REGION Network 9: Mapare elemente safety
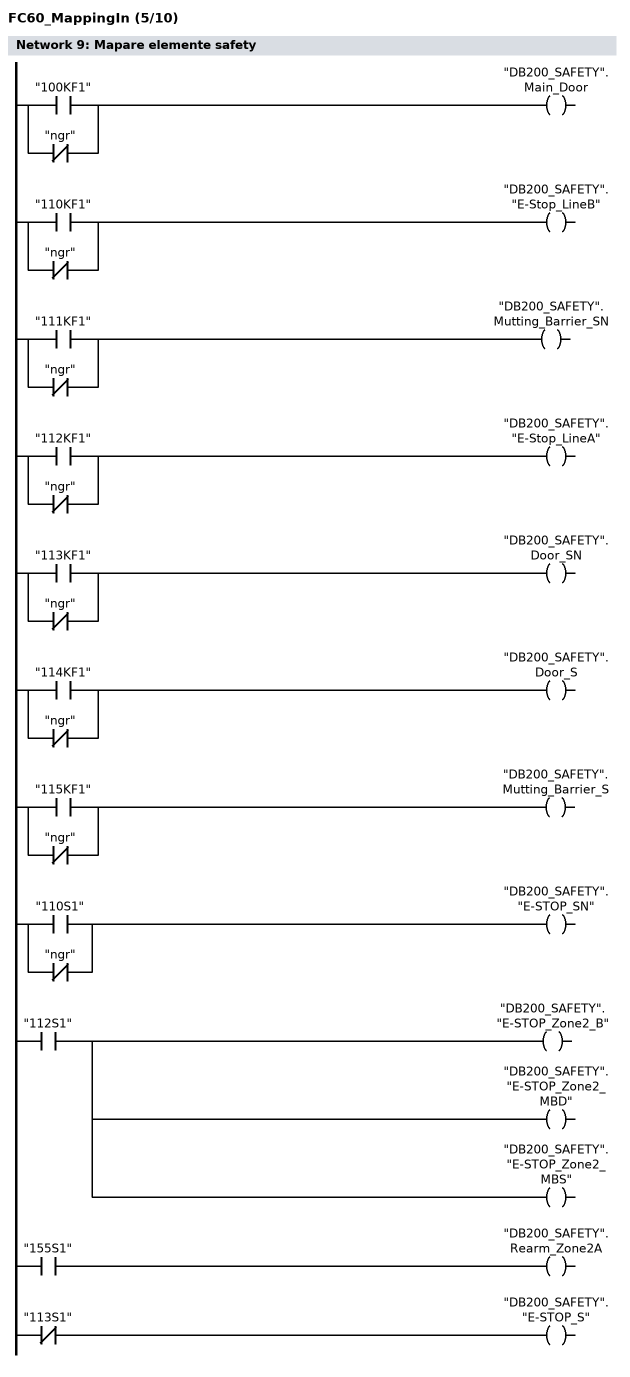
   RUNG wire#powerrail
      Contact( "100KF1" )
      wire#w1
      Coil( "DB200_SAFETY".Main_Door )
   END_RUNG
   RUNG wire#powerrail
      I_Contact( "ngr" )
   END_RUNG wire#w1
   RUNG wire#powerrail
      Contact( "110KF1" )
      wire#w2
      Coil( "DB200_SAFETY"."E-Stop_LineB" )
   END_RUNG
   RUNG wire#powerrail
      I_Contact( "ngr" )
   END_RUNG wire#w2
   RUNG wire#powerrail
      Contact( "111KF1" )
      wire#w3
      Coil( "DB200_SAFETY".Mutting_Barrier_SN )
   END_RUNG
   RUNG wire#powerrail
      I_Contact( "ngr" )
   END_RUNG wire#w3
   RUNG wire#powerrail
      Contact( "112KF1" )
      wire#w4
      Coil( "DB200_SAFETY"."E-Stop_LineA" )
   END_RUNG
   RUNG wire#powerrail
      I_Contact( "ngr" )
   END_RUNG wire#w4
   RUNG wire#powerrail
      Contact( "113KF1" )
      wire#w5
      Coil( "DB200_SAFETY".Door_SN )
   END_RUNG
   RUNG wire#powerrail
      I_Contact( "ngr" )
   END_RUNG wire#w5
   RUNG wire#powerrail
      Contact( "114KF1" )
      wire#w6
      Coil( "DB200_SAFETY".Door_S )
   END_RUNG
   RUNG wire#powerrail
      I_Contact( "ngr" )
   END_RUNG wire#w6
   RUNG wire#powerrail
      Contact( "115KF1" )
      wire#w7
      Coil( "DB200_SAFETY".Mutting_Barrier_S )
   END_RUNG
   RUNG wire#powerrail
      I_Contact( "ngr" )
   END_RUNG wire#w7
   RUNG wire#powerrail
      Contact( "110S1" )
      wire#w8
      Coil( "DB200_SAFETY"."E-STOP_SN" )
   END_RUNG
   RUNG wire#powerrail
      I_Contact( "ngr" )
   END_RUNG wire#w8
   RUNG wire#powerrail
      Contact( "112S1" )
      wire#w9
      Coil( "DB200_SAFETY"."E-STOP_Zone2_B" )
   END_RUNG
   RUNG wire#w9
      Coil( "DB200_SAFETY"."E-STOP_Zone2_MBD" )
   END_RUNG
   RUNG wire#w9
      Coil( "DB200_SAFETY"."E-STOP_Zone2_MBS" )
   END_RUNG
   RUNG wire#powerrail
      Contact( "155S1" )
      Coil( "DB200_SAFETY".Rearm_Zone2A )
   END_RUNG
   RUNG wire#powerrail
      I_Contact( "113S1" )
      Coil( "DB200_SAFETY"."E-STOP_S" )
   END_RUNG
   // the same network as SCL:
   "DB200_SAFETY".Main_Door := "100KF1" OR NOT "ngr";
   "DB200_SAFETY"."E-Stop_LineB" := "110KF1" OR NOT "ngr";
   "DB200_SAFETY".Mutting_Barrier_SN := "111KF1" OR NOT "ngr";
   "DB200_SAFETY"."E-Stop_LineA" := "112KF1" OR NOT "ngr";
   "DB200_SAFETY".Door_SN := "113KF1" OR NOT "ngr";
   "DB200_SAFETY".Door_S := "114KF1" OR NOT "ngr";
   "DB200_SAFETY".Mutting_Barrier_S := "115KF1" OR NOT "ngr";
   "DB200_SAFETY"."E-STOP_SN" := "110S1" OR NOT "ngr";
   "DB200_SAFETY"."E-STOP_Zone2_B" := "112S1";
   "DB200_SAFETY"."E-STOP_Zone2_MBD" := "112S1";
   "DB200_SAFETY"."E-STOP_Zone2_MBS" := "112S1";
   "DB200_SAFETY".Rearm_Zone2A := "155S1";
   "DB200_SAFETY"."E-STOP_S" := NOT "113S1";
END_REGION

REGION Network 10: Mapare Protectii
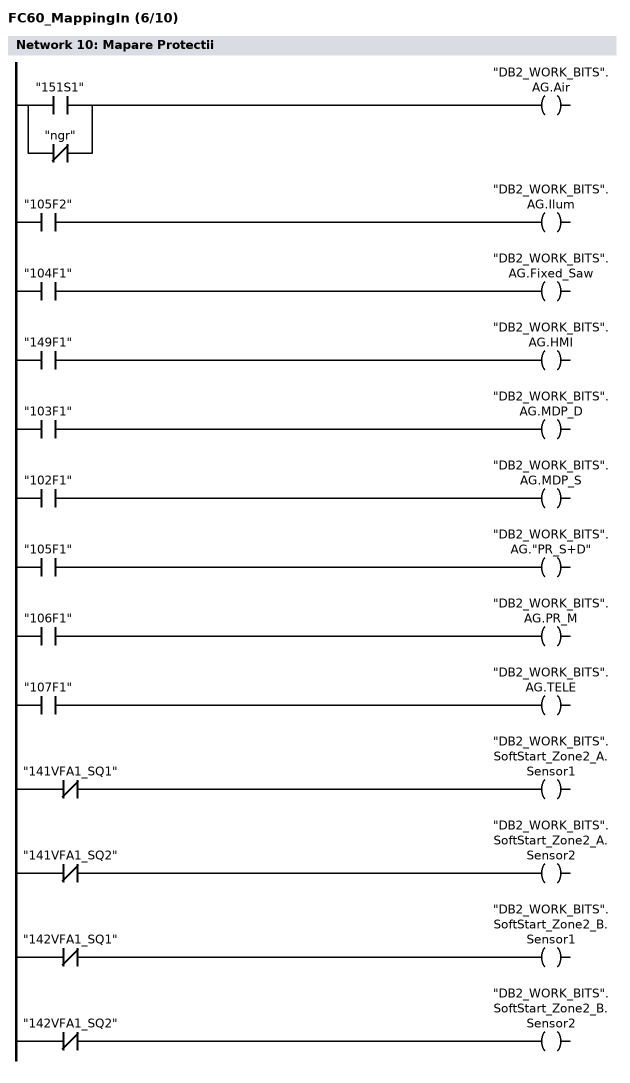
   RUNG wire#powerrail
      Contact( "151S1" )
      wire#w1
      Coil( "DB2_WORK_BITS".AG.Air )
   END_RUNG
   RUNG wire#powerrail
      I_Contact( "ngr" )
   END_RUNG wire#w1
   RUNG wire#powerrail
      Contact( "105F2" )
      Coil( "DB2_WORK_BITS".AG.Ilum )
   END_RUNG
   RUNG wire#powerrail
      Contact( "104F1" )
      Coil( "DB2_WORK_BITS".AG.Fixed_Saw )
   END_RUNG
   RUNG wire#powerrail
      Contact( "149F1" )
      Coil( "DB2_WORK_BITS".AG.HMI )
   END_RUNG
   RUNG wire#powerrail
      Contact( "103F1" )
      Coil( "DB2_WORK_BITS".AG.MDP_D )
   END_RUNG
   RUNG wire#powerrail
      Contact( "102F1" )
      Coil( "DB2_WORK_BITS".AG.MDP_S )
   END_RUNG
   RUNG wire#powerrail
      Contact( "105F1" )
      Coil( "DB2_WORK_BITS".AG."PR_S+D" )
   END_RUNG
   RUNG wire#powerrail
      Contact( "106F1" )
      Coil( "DB2_WORK_BITS".AG.PR_M )
   END_RUNG
   RUNG wire#powerrail
      Contact( "107F1" )
      Coil( "DB2_WORK_BITS".AG.TELE )
   END_RUNG
   RUNG wire#powerrail
      I_Contact( "141VFA1_SQ1" )
      Coil( "DB2_WORK_BITS".SoftStart_Zone2_A.Sensor1 )
   END_RUNG
   RUNG wire#powerrail
      I_Contact( "141VFA1_SQ2" )
      Coil( "DB2_WORK_BITS".SoftStart_Zone2_A.Sensor2 )
   END_RUNG
   RUNG wire#powerrail
      I_Contact( "142VFA1_SQ1" )
      Coil( "DB2_WORK_BITS".SoftStart_Zone2_B.Sensor1 )
   END_RUNG
   RUNG wire#powerrail
      I_Contact( "142VFA1_SQ2" )
      Coil( "DB2_WORK_BITS".SoftStart_Zone2_B.Sensor2 )
   END_RUNG
   // the same network as SCL:
   "DB2_WORK_BITS".AG.Air := "151S1" OR NOT "ngr";
   "DB2_WORK_BITS".AG.Ilum := "105F2";
   "DB2_WORK_BITS".AG.Fixed_Saw := "104F1";
   "DB2_WORK_BITS".AG.HMI := "149F1";
   "DB2_WORK_BITS".AG.MDP_D := "103F1";
   "DB2_WORK_BITS".AG.MDP_S := "102F1";
   "DB2_WORK_BITS".AG."PR_S+D" := "105F1";
   "DB2_WORK_BITS".AG.PR_M := "106F1";
   "DB2_WORK_BITS".AG.TELE := "107F1";
   "DB2_WORK_BITS".SoftStart_Zone2_A.Sensor1 := NOT "141VFA1_SQ1";
   "DB2_WORK_BITS".SoftStart_Zone2_A.Sensor2 := NOT "141VFA1_SQ2";
   "DB2_WORK_BITS".SoftStart_Zone2_B.Sensor1 := NOT "142VFA1_SQ1";
   "DB2_WORK_BITS".SoftStart_Zone2_B.Sensor2 := NOT "142VFA1_SQ2";
END_REGION

REGION Network 11: Stacker_Nou Conveior 1
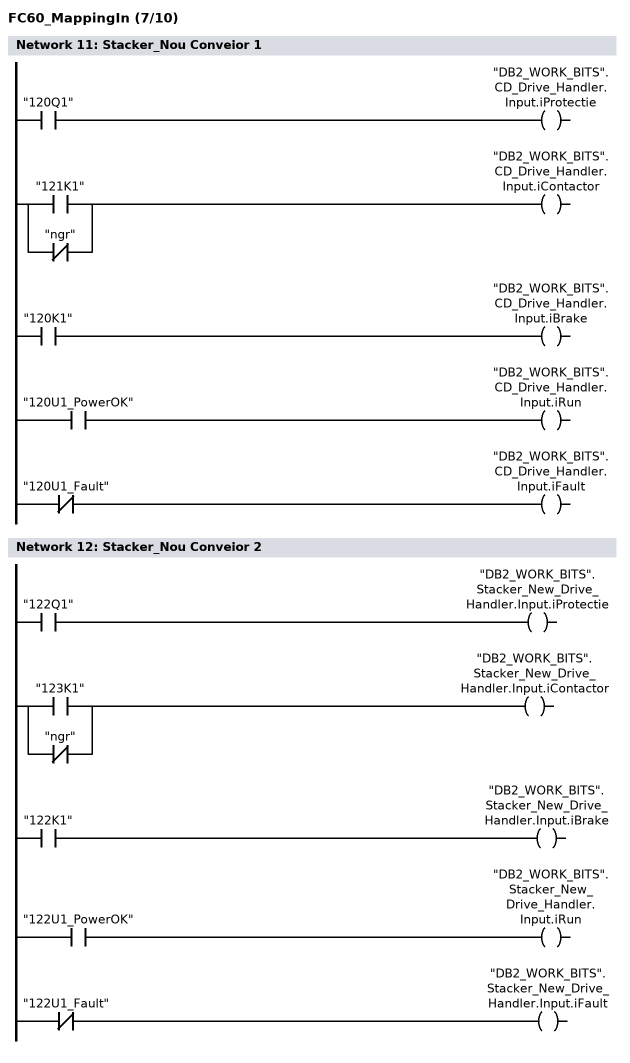
   RUNG wire#powerrail
      Contact( "120Q1" )
      Coil( "DB2_WORK_BITS".CD_Drive_Handler.Input.iProtectie )
   END_RUNG
   RUNG wire#powerrail
      Contact( "121K1" )
      wire#w1
      Coil( "DB2_WORK_BITS".CD_Drive_Handler.Input.iContactor )
   END_RUNG
   RUNG wire#powerrail
      I_Contact( "ngr" )
   END_RUNG wire#w1
   RUNG wire#powerrail
      Contact( "120K1" )
      Coil( "DB2_WORK_BITS".CD_Drive_Handler.Input.iBrake )
   END_RUNG
   RUNG wire#powerrail
      Contact( "120U1_PowerOK" )
      Coil( "DB2_WORK_BITS".CD_Drive_Handler.Input.iRun )
   END_RUNG
   RUNG wire#powerrail
      I_Contact( "120U1_Fault" )
      Coil( "DB2_WORK_BITS".CD_Drive_Handler.Input.iFault )
   END_RUNG
   // the same network as SCL:
   "DB2_WORK_BITS".CD_Drive_Handler.Input.iProtectie := "120Q1";
   "DB2_WORK_BITS".CD_Drive_Handler.Input.iContactor := "121K1" OR NOT "ngr";
   "DB2_WORK_BITS".CD_Drive_Handler.Input.iBrake := "120K1";
   "DB2_WORK_BITS".CD_Drive_Handler.Input.iRun := "120U1_PowerOK";
   "DB2_WORK_BITS".CD_Drive_Handler.Input.iFault := NOT "120U1_Fault";
END_REGION

REGION Network 12: Stacker_Nou Conveior 2
   RUNG wire#powerrail
      Contact( "122Q1" )
      Coil( "DB2_WORK_BITS".Stacker_New_Drive_Handler.Input.iProtectie )
   END_RUNG
   RUNG wire#powerrail
      Contact( "123K1" )
      wire#w1
      Coil( "DB2_WORK_BITS".Stacker_New_Drive_Handler.Input.iContactor )
   END_RUNG
   RUNG wire#powerrail
      I_Contact( "ngr" )
   END_RUNG wire#w1
   RUNG wire#powerrail
      Contact( "122K1" )
      Coil( "DB2_WORK_BITS".Stacker_New_Drive_Handler.Input.iBrake )
   END_RUNG
   RUNG wire#powerrail
      Contact( "122U1_PowerOK" )
      Coil( "DB2_WORK_BITS".Stacker_New_Drive_Handler.Input.iRun )
   END_RUNG
   RUNG wire#powerrail
      I_Contact( "122U1_Fault" )
      Coil( "DB2_WORK_BITS".Stacker_New_Drive_Handler.Input.iFault )
   END_RUNG
   // the same network as SCL:
   "DB2_WORK_BITS".Stacker_New_Drive_Handler.Input.iProtectie := "122Q1";
   "DB2_WORK_BITS".Stacker_New_Drive_Handler.Input.iContactor := "123K1" OR NOT "ngr";
   "DB2_WORK_BITS".Stacker_New_Drive_Handler.Input.iBrake := "122K1";
   "DB2_WORK_BITS".Stacker_New_Drive_Handler.Input.iRun := "122U1_PowerOK";
   "DB2_WORK_BITS".Stacker_New_Drive_Handler.Input.iFault := NOT "122U1_Fault";
END_REGION

REGION Network 13: Zona B
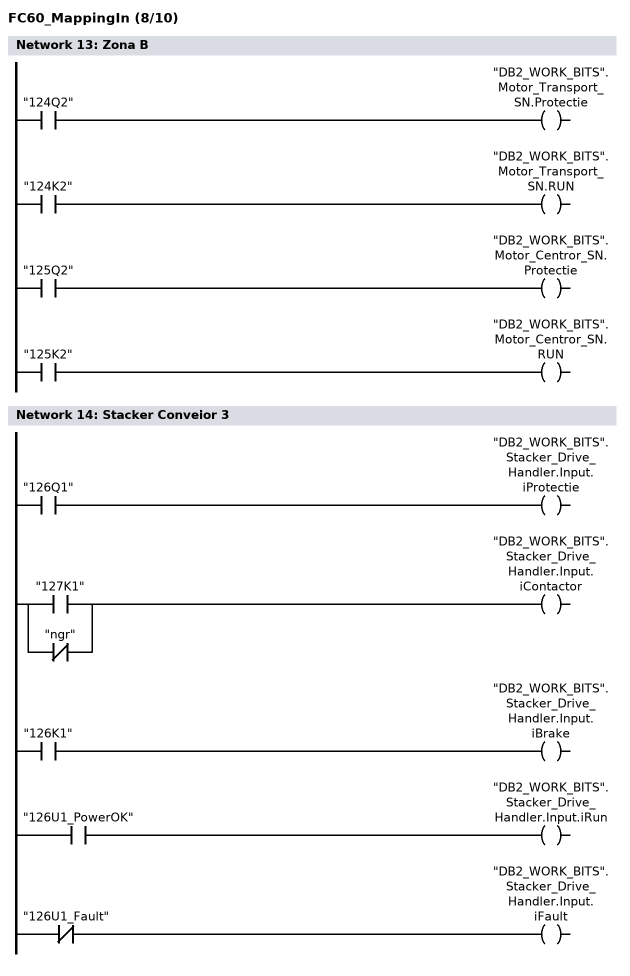
   RUNG wire#powerrail
      Contact( "124Q2" )
      Coil( "DB2_WORK_BITS".Motor_Transport_SN.Protectie )
   END_RUNG
   RUNG wire#powerrail
      Contact( "124K2" )
      Coil( "DB2_WORK_BITS".Motor_Transport_SN.RUN )
   END_RUNG
   RUNG wire#powerrail
      Contact( "125Q2" )
      Coil( "DB2_WORK_BITS".Motor_Centror_SN.Protectie )
   END_RUNG
   RUNG wire#powerrail
      Contact( "125K2" )
      Coil( "DB2_WORK_BITS".Motor_Centror_SN.RUN )
   END_RUNG
   // the same network as SCL:
   "DB2_WORK_BITS".Motor_Transport_SN.Protectie := "124Q2";
   "DB2_WORK_BITS".Motor_Transport_SN.RUN := "124K2";
   "DB2_WORK_BITS".Motor_Centror_SN.Protectie := "125Q2";
   "DB2_WORK_BITS".Motor_Centror_SN.RUN := "125K2";
END_REGION

REGION Network 14: Stacker Conveior 3
   RUNG wire#powerrail
      Contact( "126Q1" )
      Coil( "DB2_WORK_BITS".Stacker_Drive_Handler.Input.iProtectie )
   END_RUNG
   RUNG wire#powerrail
      Contact( "127K1" )
      wire#w1
      Coil( "DB2_WORK_BITS".Stacker_Drive_Handler.Input.iContactor )
   END_RUNG
   RUNG wire#powerrail
      I_Contact( "ngr" )
   END_RUNG wire#w1
   RUNG wire#powerrail
      Contact( "126K1" )
      Coil( "DB2_WORK_BITS".Stacker_Drive_Handler.Input.iBrake )
   END_RUNG
   RUNG wire#powerrail
      Contact( "126U1_PowerOK" )
      Coil( "DB2_WORK_BITS".Stacker_Drive_Handler.Input.iRun )
   END_RUNG
   RUNG wire#powerrail
      I_Contact( "126U1_Fault" )
      Coil( "DB2_WORK_BITS".Stacker_Drive_Handler.Input.iFault )
   END_RUNG
   // the same network as SCL:
   "DB2_WORK_BITS".Stacker_Drive_Handler.Input.iProtectie := "126Q1";
   "DB2_WORK_BITS".Stacker_Drive_Handler.Input.iContactor := "127K1" OR NOT "ngr";
   "DB2_WORK_BITS".Stacker_Drive_Handler.Input.iBrake := "126K1";
   "DB2_WORK_BITS".Stacker_Drive_Handler.Input.iRun := "126U1_PowerOK";
   "DB2_WORK_BITS".Stacker_Drive_Handler.Input.iFault := NOT "126U1_Fault";
END_REGION

REGION Network 15: Stacker Conveior 4
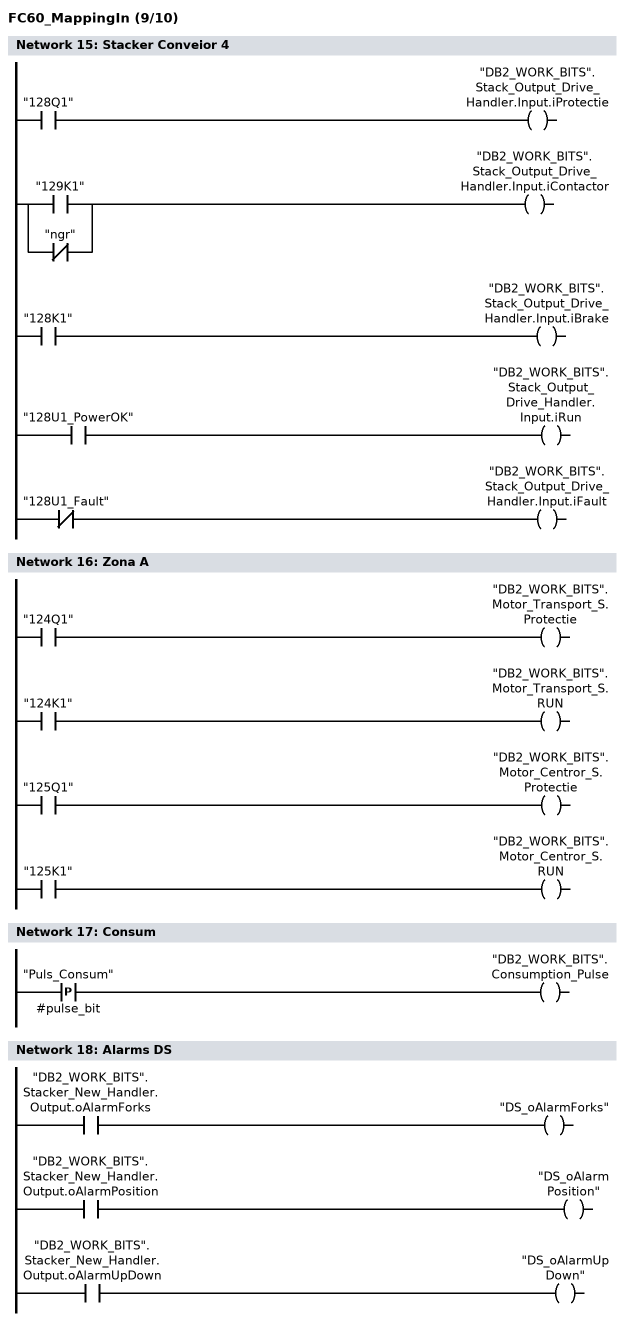
   RUNG wire#powerrail
      Contact( "128Q1" )
      Coil( "DB2_WORK_BITS".Stack_Output_Drive_Handler.Input.iProtectie )
   END_RUNG
   RUNG wire#powerrail
      Contact( "129K1" )
      wire#w1
      Coil( "DB2_WORK_BITS".Stack_Output_Drive_Handler.Input.iContactor )
   END_RUNG
   RUNG wire#powerrail
      I_Contact( "ngr" )
   END_RUNG wire#w1
   RUNG wire#powerrail
      Contact( "128K1" )
      Coil( "DB2_WORK_BITS".Stack_Output_Drive_Handler.Input.iBrake )
   END_RUNG
   RUNG wire#powerrail
      Contact( "128U1_PowerOK" )
      Coil( "DB2_WORK_BITS".Stack_Output_Drive_Handler.Input.iRun )
   END_RUNG
   RUNG wire#powerrail
      I_Contact( "128U1_Fault" )
      Coil( "DB2_WORK_BITS".Stack_Output_Drive_Handler.Input.iFault )
   END_RUNG
   // the same network as SCL:
   "DB2_WORK_BITS".Stack_Output_Drive_Handler.Input.iProtectie := "128Q1";
   "DB2_WORK_BITS".Stack_Output_Drive_Handler.Input.iContactor := "129K1" OR NOT "ngr";
   "DB2_WORK_BITS".Stack_Output_Drive_Handler.Input.iBrake := "128K1";
   "DB2_WORK_BITS".Stack_Output_Drive_Handler.Input.iRun := "128U1_PowerOK";
   "DB2_WORK_BITS".Stack_Output_Drive_Handler.Input.iFault := NOT "128U1_Fault";
END_REGION

REGION Network 16: Zona A
   RUNG wire#powerrail
      Contact( "124Q1" )
      Coil( "DB2_WORK_BITS".Motor_Transport_S.Protectie )
   END_RUNG
   RUNG wire#powerrail
      Contact( "124K1" )
      Coil( "DB2_WORK_BITS".Motor_Transport_S.RUN )
   END_RUNG
   RUNG wire#powerrail
      Contact( "125Q1" )
      Coil( "DB2_WORK_BITS".Motor_Centror_S.Protectie )
   END_RUNG
   RUNG wire#powerrail
      Contact( "125K1" )
      Coil( "DB2_WORK_BITS".Motor_Centror_S.RUN )
   END_RUNG
   // the same network as SCL:
   "DB2_WORK_BITS".Motor_Transport_S.Protectie := "124Q1";
   "DB2_WORK_BITS".Motor_Transport_S.RUN := "124K1";
   "DB2_WORK_BITS".Motor_Centror_S.Protectie := "125Q1";
   "DB2_WORK_BITS".Motor_Centror_S.RUN := "125K1";
END_REGION

REGION Network 17: Consum
   RUNG wire#powerrail
      P_Contact(operand := "Puls_Consum", bit := #pulse_bit)
      Coil( "DB2_WORK_BITS".Consumption_Pulse )
   END_RUNG
   // the same network as SCL:
   #_w1 := "Puls_Consum" AND NOT #pulse_bit;   // rising edge of "Puls_Consum"
   #pulse_bit := "Puls_Consum";
   "DB2_WORK_BITS".Consumption_Pulse := #_w1;
END_REGION

REGION Network 18: Alarms DS
   RUNG wire#powerrail
      Contact( "DB2_WORK_BITS".Stacker_New_Handler.Output.oAlarmForks )
      Coil( "DS_oAlarmForks" )
   END_RUNG
   RUNG wire#powerrail
      Contact( "DB2_WORK_BITS".Stacker_New_Handler.Output.oAlarmPosition )
      Coil( "DS_oAlarmPosition" )
   END_RUNG
   RUNG wire#powerrail
      Contact( "DB2_WORK_BITS".Stacker_New_Handler.Output.oAlarmUpDown )
      Coil( "DS_oAlarmUpDown" )
   END_RUNG
   // the same network as SCL:
   "DS_oAlarmForks" := "DB2_WORK_BITS".Stacker_New_Handler.Output.oAlarmForks;
   "DS_oAlarmPosition" := "DB2_WORK_BITS".Stacker_New_Handler.Output.oAlarmPosition;
   "DS_oAlarmUpDown" := "DB2_WORK_BITS".Stacker_New_Handler.Output.oAlarmUpDown;
END_REGION

REGION Network 19: Alarms S
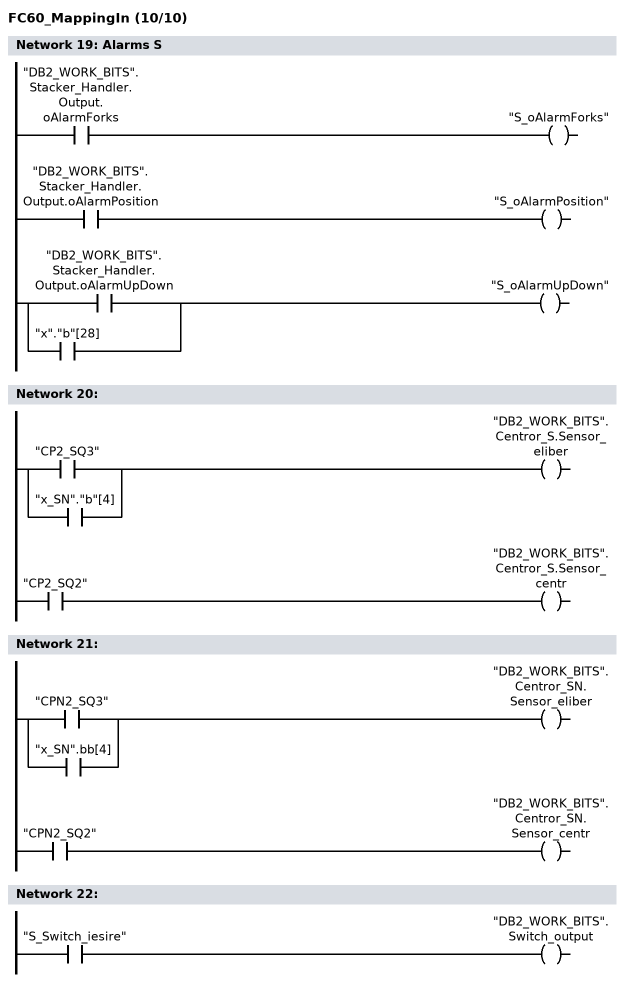
   RUNG wire#powerrail
      Contact( "DB2_WORK_BITS".Stacker_Handler.Output.oAlarmForks )
      Coil( "S_oAlarmForks" )
   END_RUNG
   RUNG wire#powerrail
      Contact( "DB2_WORK_BITS".Stacker_Handler.Output.oAlarmPosition )
      Coil( "S_oAlarmPosition" )
   END_RUNG
   RUNG wire#powerrail
      Contact( "DB2_WORK_BITS".Stacker_Handler.Output.oAlarmUpDown )
      wire#w1
      Coil( "S_oAlarmUpDown" )
   END_RUNG
   RUNG wire#powerrail
      Contact( "x"."b"[28] )
   END_RUNG wire#w1
   // the same network as SCL:
   "S_oAlarmForks" := "DB2_WORK_BITS".Stacker_Handler.Output.oAlarmForks;
   "S_oAlarmPosition" := "DB2_WORK_BITS".Stacker_Handler.Output.oAlarmPosition;
   "S_oAlarmUpDown" := "DB2_WORK_BITS".Stacker_Handler.Output.oAlarmUpDown OR "x"."b"[28];
END_REGION

REGION Network 20
   RUNG wire#powerrail
      Contact( "CP2_SQ3" )
      wire#w1
      Coil( "DB2_WORK_BITS".Centror_S.Sensor_eliber )
   END_RUNG
   RUNG wire#powerrail
      Contact( "x_SN"."b"[4] )
   END_RUNG wire#w1
   RUNG wire#powerrail
      Contact( "CP2_SQ2" )
      Coil( "DB2_WORK_BITS".Centror_S.Sensor_centr )
   END_RUNG
   // the same network as SCL:
   "DB2_WORK_BITS".Centror_S.Sensor_eliber := "CP2_SQ3" OR "x_SN"."b"[4];
   "DB2_WORK_BITS".Centror_S.Sensor_centr := "CP2_SQ2";
END_REGION

REGION Network 21
   RUNG wire#powerrail
      Contact( "CPN2_SQ3" )
      wire#w1
      Coil( "DB2_WORK_BITS".Centror_SN.Sensor_eliber )
   END_RUNG
   RUNG wire#powerrail
      Contact( "x_SN".bb[4] )
   END_RUNG wire#w1
   RUNG wire#powerrail
      Contact( "CPN2_SQ2" )
      Coil( "DB2_WORK_BITS".Centror_SN.Sensor_centr )
   END_RUNG
   // the same network as SCL:
   "DB2_WORK_BITS".Centror_SN.Sensor_eliber := "CPN2_SQ3" OR "x_SN".bb[4];
   "DB2_WORK_BITS".Centror_SN.Sensor_centr := "CPN2_SQ2";
END_REGION

REGION Network 22
   RUNG wire#powerrail
      Contact( "S_Switch_iesire" )
      Coil( "DB2_WORK_BITS".Switch_output )
   END_RUNG
   // the same network as SCL:
   "DB2_WORK_BITS".Switch_output := "S_Switch_iesire";
END_REGION
END_FUNCTION

FUNCTION "FC3_FAULTS" : Void   // FC3, LAD
{ S7_Optimized_Access := 'TRUE' }
VERSION : 0.1
   VAR_TEMP
      ctrlLoop : Bool;
      orResult : Bool;
      NoAlmStop : Bool;
      NoAlmAny : Bool;
      SN_NoAlmAny : Bool;
   END_VAR
   VAR_TEMP   // added for the SCL form of the ladder/FBD networks
      _w1 : Bool;
   END_VAR
BEGIN

REGION Network 1: rst
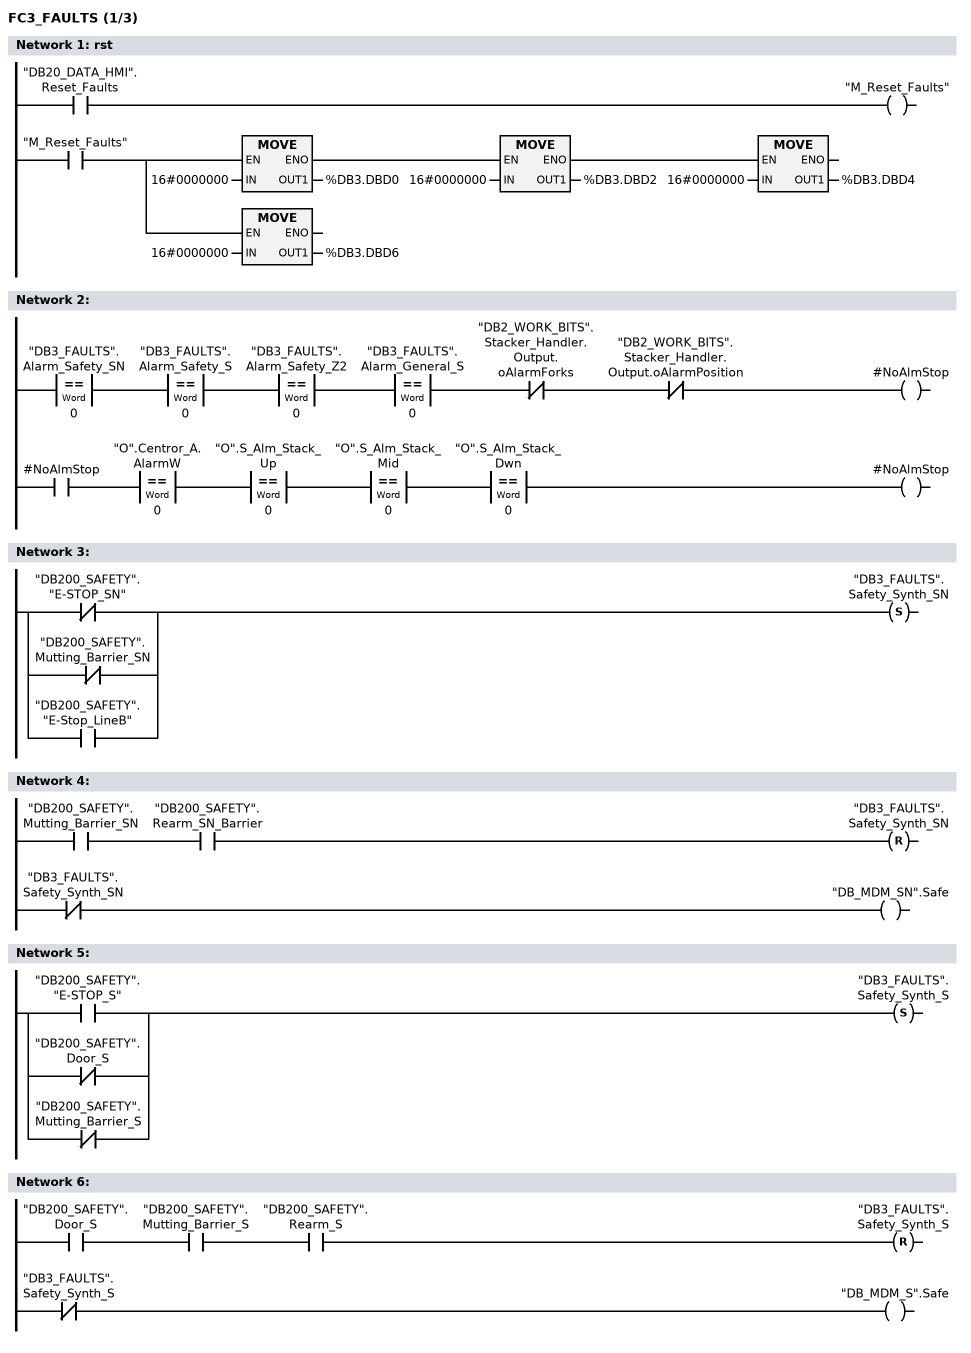
   RUNG wire#powerrail
      Contact( "DB20_DATA_HMI".Reset_Faults )
      Coil( "M_Reset_Faults" )
   END_RUNG
   RUNG wire#powerrail
      Contact( "M_Reset_Faults" )
      wire#w1
      Move(in := 16#0000000, out1 => %DB3.DBD0)
      Move(in := 16#0000000, out1 => %DB3.DBD2)
      Move(in := 16#0000000, out1 => %DB3.DBD4)
   END_RUNG
   RUNG wire#w1
      Move(in := 16#0000000, out1 => %DB3.DBD6)
   END_RUNG
   // the same network as SCL:
   "M_Reset_Faults" := "DB20_DATA_HMI".Reset_Faults;
   IF "M_Reset_Faults" THEN
       %DB3.DBD0 := 16#0000000;
       %DB3.DBD2 := 16#0000000;
       %DB3.DBD4 := 16#0000000;
       %DB3.DBD6 := 16#0000000;
   END_IF;
END_REGION

REGION Network 2
   RUNG wire#powerrail
      { S7_Templates := "SrcType := Word" } EQ_Contact(in1 := "DB3_FAULTS".Alarm_Safety_SN, in2 := 0)
      { S7_Templates := "SrcType := Word" } EQ_Contact(in1 := "DB3_FAULTS".Alarm_Safety_S, in2 := 0)
      { S7_Templates := "SrcType := Word" } EQ_Contact(in1 := "DB3_FAULTS".Alarm_Safety_Z2, in2 := 0)
      { S7_Templates := "SrcType := Word" } EQ_Contact(in1 := "DB3_FAULTS".Alarm_General_S, in2 := 0)
      I_Contact( "DB2_WORK_BITS".Stacker_Handler.Output.oAlarmForks )
      I_Contact( "DB2_WORK_BITS".Stacker_Handler.Output.oAlarmPosition )
      Coil( #NoAlmStop )
   END_RUNG
   RUNG wire#powerrail
      Contact( #NoAlmStop )
      { S7_Templates := "SrcType := Word" } EQ_Contact(in1 := "O".Centror_A.AlarmW, in2 := 0)
      { S7_Templates := "SrcType := Word" } EQ_Contact(in1 := "O".S_Alm_Stack_Up, in2 := 0)
      { S7_Templates := "SrcType := Word" } EQ_Contact(in1 := "O".S_Alm_Stack_Mid, in2 := 0)
      { S7_Templates := "SrcType := Word" } EQ_Contact(in1 := "O".S_Alm_Stack_Dwn, in2 := 0)
      Coil( #NoAlmStop )
   END_RUNG
   // the same network as SCL:
   #NoAlmStop := ("DB3_FAULTS".Alarm_Safety_SN = 0) AND ("DB3_FAULTS".Alarm_Safety_S = 0) AND ("DB3_FAULTS".Alarm_Safety_Z2 = 0) AND ("DB3_FAULTS".Alarm_General_S = 0) AND NOT "DB2_WORK_BITS".Stacker_Handler.Output.oAlarmForks AND NOT "DB2_WORK_BITS".Stacker_Handler.Output.oAlarmPosition;
   #NoAlmStop := #NoAlmStop AND ("O".Centror_A.AlarmW = 0) AND ("O".S_Alm_Stack_Up = 0) AND ("O".S_Alm_Stack_Mid = 0) AND ("O".S_Alm_Stack_Dwn = 0);
END_REGION

REGION Network 3
   RUNG wire#powerrail
      I_Contact( "DB200_SAFETY"."E-STOP_SN" )
      wire#w1
      S_Coil( "DB3_FAULTS".Safety_Synth_SN )
   END_RUNG
   RUNG wire#powerrail
      I_Contact( "DB200_SAFETY".Mutting_Barrier_SN )
   END_RUNG wire#w1
   RUNG wire#powerrail
      Contact( "DB200_SAFETY"."E-Stop_LineB" )
   END_RUNG wire#w1
   // the same network as SCL:
   IF NOT "DB200_SAFETY"."E-STOP_SN" OR NOT "DB200_SAFETY".Mutting_Barrier_SN OR "DB200_SAFETY"."E-Stop_LineB" THEN
       "DB3_FAULTS".Safety_Synth_SN := TRUE;
   END_IF;
END_REGION

REGION Network 4
   RUNG wire#powerrail
      Contact( "DB200_SAFETY".Mutting_Barrier_SN )
      Contact( "DB200_SAFETY".Rearm_SN_Barrier )
      R_Coil( "DB3_FAULTS".Safety_Synth_SN )
   END_RUNG
   RUNG wire#powerrail
      I_Contact( "DB3_FAULTS".Safety_Synth_SN )
      Coil( "DB_MDM_SN".Safe )
   END_RUNG
   // the same network as SCL:
   IF "DB200_SAFETY".Mutting_Barrier_SN AND "DB200_SAFETY".Rearm_SN_Barrier THEN
       "DB3_FAULTS".Safety_Synth_SN := FALSE;
   END_IF;
   "DB_MDM_SN".Safe := NOT "DB3_FAULTS".Safety_Synth_SN;
END_REGION

REGION Network 5
   RUNG wire#powerrail
      Contact( "DB200_SAFETY"."E-STOP_S" )
      wire#w1
      S_Coil( "DB3_FAULTS".Safety_Synth_S )
   END_RUNG
   RUNG wire#powerrail
      I_Contact( "DB200_SAFETY".Door_S )
   END_RUNG wire#w1
   RUNG wire#powerrail
      I_Contact( "DB200_SAFETY".Mutting_Barrier_S )
   END_RUNG wire#w1
   // the same network as SCL:
   IF "DB200_SAFETY"."E-STOP_S" OR NOT "DB200_SAFETY".Door_S OR NOT "DB200_SAFETY".Mutting_Barrier_S THEN
       "DB3_FAULTS".Safety_Synth_S := TRUE;
   END_IF;
END_REGION

REGION Network 6
   RUNG wire#powerrail
      Contact( "DB200_SAFETY".Door_S )
      Contact( "DB200_SAFETY".Mutting_Barrier_S )
      Contact( "DB200_SAFETY".Rearm_S )
      R_Coil( "DB3_FAULTS".Safety_Synth_S )
   END_RUNG
   RUNG wire#powerrail
      I_Contact( "DB3_FAULTS".Safety_Synth_S )
      Coil( "DB_MDM_S".Safe )
   END_RUNG
   // the same network as SCL:
   IF "DB200_SAFETY".Door_S AND "DB200_SAFETY".Mutting_Barrier_S AND "DB200_SAFETY".Rearm_S THEN
       "DB3_FAULTS".Safety_Synth_S := FALSE;
   END_IF;
   "DB_MDM_S".Safe := NOT "DB3_FAULTS".Safety_Synth_S;
END_REGION

REGION Network 7
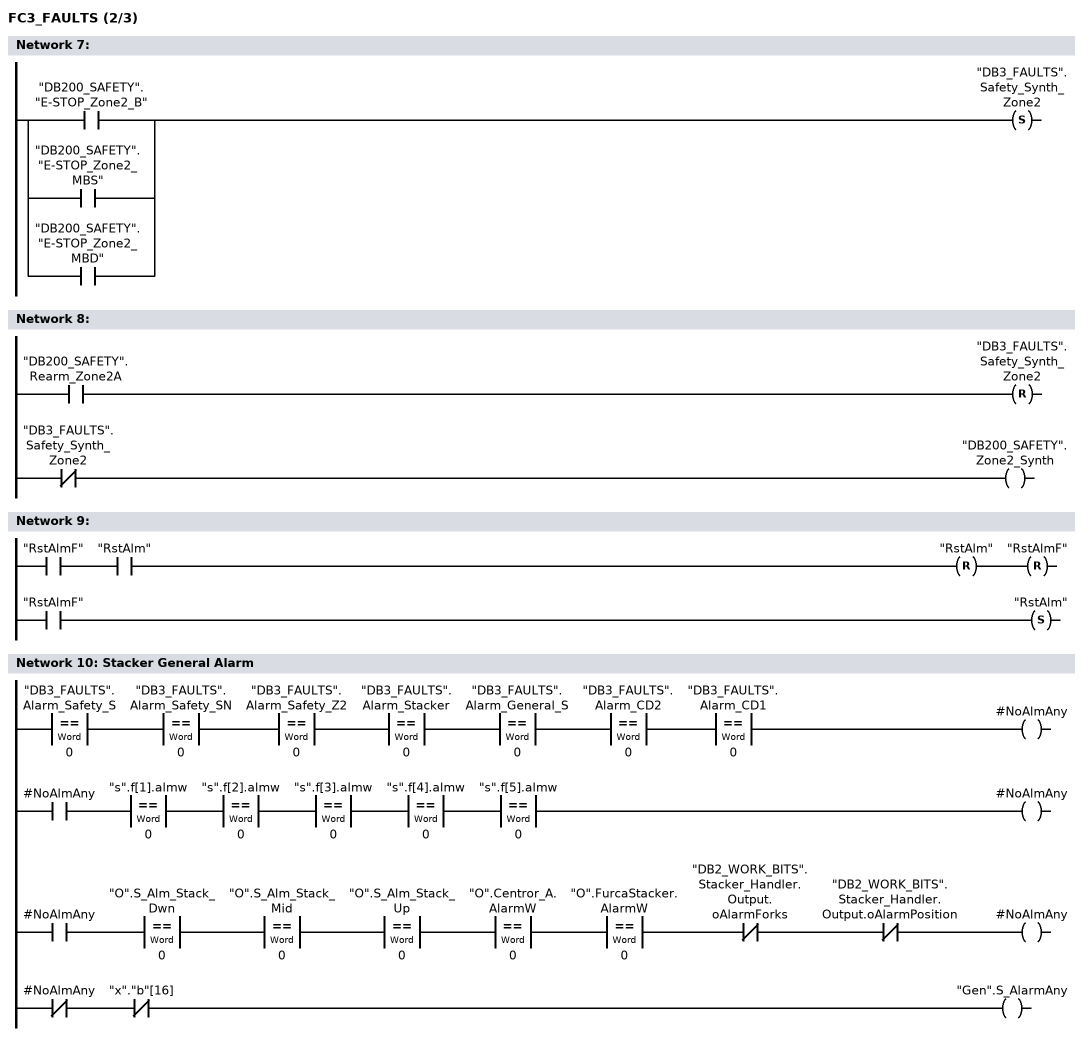
   RUNG wire#powerrail
      Contact( "DB200_SAFETY"."E-STOP_Zone2_B" )
      wire#w1
      S_Coil( "DB3_FAULTS".Safety_Synth_Zone2 )
   END_RUNG
   RUNG wire#powerrail
      Contact( "DB200_SAFETY"."E-STOP_Zone2_MBS" )
   END_RUNG wire#w1
   RUNG wire#powerrail
      Contact( "DB200_SAFETY"."E-STOP_Zone2_MBD" )
   END_RUNG wire#w1
   // the same network as SCL:
   IF "DB200_SAFETY"."E-STOP_Zone2_B" OR "DB200_SAFETY"."E-STOP_Zone2_MBS" OR "DB200_SAFETY"."E-STOP_Zone2_MBD" THEN
       "DB3_FAULTS".Safety_Synth_Zone2 := TRUE;
   END_IF;
END_REGION

REGION Network 8
   RUNG wire#powerrail
      Contact( "DB200_SAFETY".Rearm_Zone2A )
      R_Coil( "DB3_FAULTS".Safety_Synth_Zone2 )
   END_RUNG
   RUNG wire#powerrail
      I_Contact( "DB3_FAULTS".Safety_Synth_Zone2 )
      Coil( "DB200_SAFETY".Zone2_Synth )
   END_RUNG
   // the same network as SCL:
   IF "DB200_SAFETY".Rearm_Zone2A THEN "DB3_FAULTS".Safety_Synth_Zone2 := FALSE; END_IF;
   "DB200_SAFETY".Zone2_Synth := NOT "DB3_FAULTS".Safety_Synth_Zone2;
END_REGION

REGION Network 9
   RUNG wire#powerrail
      Contact( "RstAlmF" )
      Contact( "RstAlm" )
      R_Coil( "RstAlm" )
      R_Coil( "RstAlmF" )
   END_RUNG
   RUNG wire#powerrail
      Contact( "RstAlmF" )
      S_Coil( "RstAlm" )
   END_RUNG
   // the same network as SCL:
   #_w1 := "RstAlmF" AND "RstAlm";
   IF #_w1 THEN
       "RstAlm" := FALSE;
       "RstAlmF" := FALSE;
   END_IF;
   IF "RstAlmF" THEN "RstAlm" := TRUE; END_IF;
END_REGION
